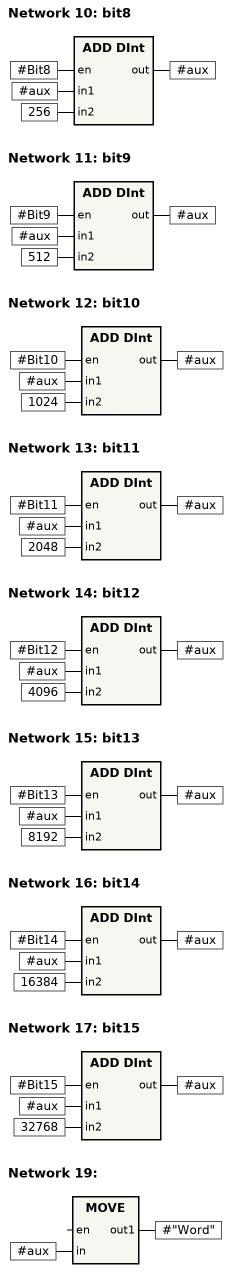
   IF #Bit8 THEN #aux := #aux + 256; END_IF;
END_REGION

REGION Network 11: bit9
   // Addiere Bit 9 zur Hilfsvariable "aux".
   // ***************************************************************************
   // Add Bit 9 to the auxiliary variable "aux".
   IF #Bit9 THEN #aux := #aux + 512; END_IF;
END_REGION

REGION Network 12: bit10
   // Addiere Bit 10 zur Hilfsvariable "aux".
   // ***************************************************************************
   // Add Bit 10 to the auxiliary variable "aux".
   IF #Bit10 THEN #aux := #aux + 1024; END_IF;
END_REGION

REGION Network 13: bit11
   // Addiere Bit 11 zur Hilfsvariable "aux".
   // ***************************************************************************
   // Add Bit 11 to the auxiliary variable "aux".
   IF #Bit11 THEN #aux := #aux + 2048; END_IF;
END_REGION

REGION Network 14: bit12
   // Addiere Bit 12 zur Hilfsvariable "aux".
   // ***************************************************************************
   // Add Bit 12 to the auxiliary variable "aux".
   IF #Bit12 THEN #aux := #aux + 4096; END_IF;
END_REGION

REGION Network 15: bit13
   // Addiere Bit 13 zur Hilfsvariable "aux".
   // ***************************************************************************
   // Add Bit 13 to the auxiliary variable "aux".
   IF #Bit13 THEN #aux := #aux + 8192; END_IF;
END_REGION

REGION Network 16: bit14
   // Addiere Bit 14 zur Hilfsvariable "aux".
   // ***************************************************************************
   // Add Bit 14 to the auxiliary variable "aux".
   IF #Bit14 THEN #aux := #aux + 16384; END_IF;
END_REGION

REGION Network 17: bit15
   // Addiere Bit 15 zur Hilfsvariable "aux".
   // ***************************************************************************
   // Add Bit 15 to the auxiliary variable "aux".
   IF #Bit15 THEN #aux := #aux + 32768; END_IF;
END_REGION

REGION Network 18: Word
   // Der Wert der Variablen "aux" wird  vom Datentyp "UInt" zum Datentyp "Word" konvertiert und der Ausgangsvariablen "Word" übergeben.
   // ***************************************************************************
   // The value of the variable "aux" will convert from type of data "UInt" to type of data "Word" and transfered to the output variable "Word".
END_REGION

REGION Network 19
   #"Word" := #aux;
END_REGION
END_FUNCTION

// folder: 60 - 69 Alarm & Satus Handling

FUNCTION "60_Alarms" : Void   // FC60, LAD
TITLE = Alarm Processing
{ S7_Optimized_Access := 'TRUE' }
AUTHOR : JRS
VERSION : 0.1
// To determine alarm conditions
   VAR_TEMP   // added for the SCL form of the ladder/FBD networks
      _w1 : Bool;
      _w2 : Bool;
   END_VAR
BEGIN

REGION Network 1: DB60 DBX0.0 = Master PLC Heart Beat Missing
   // BC_ALARM_WORD_01_BIT_0
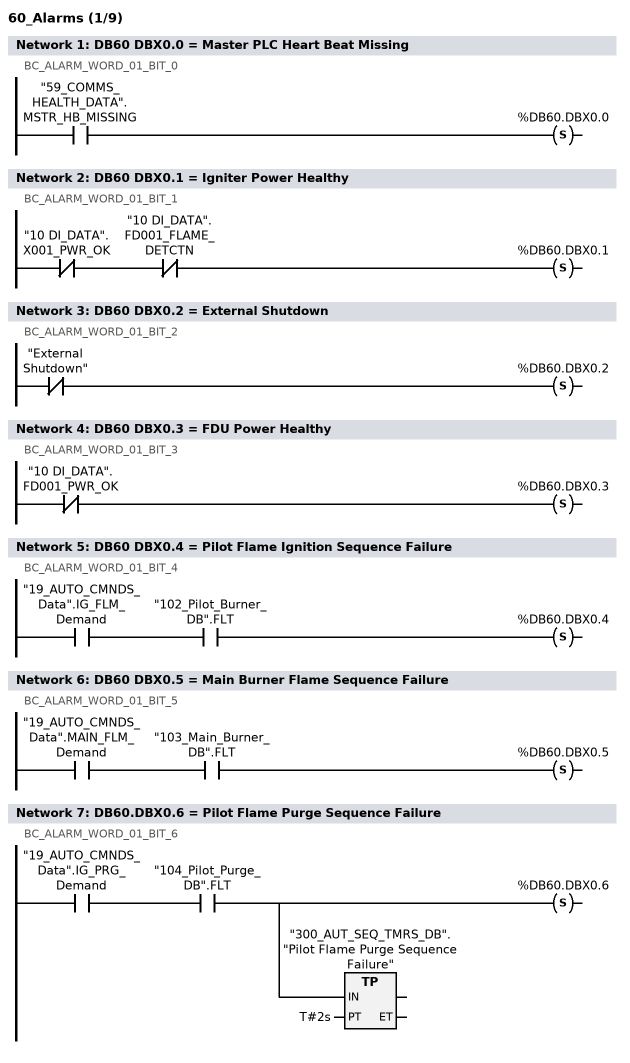
   RUNG wire#powerrail
      Contact( "59_COMMS_HEALTH_DATA".MSTR_HB_MISSING )
      S_Coil( %DB60.DBX0.0 )
   END_RUNG
   // the same network as SCL:
   IF "59_COMMS_HEALTH_DATA".MSTR_HB_MISSING THEN %DB60.DBX0.0 := TRUE; END_IF;
END_REGION

REGION Network 2: DB60 DBX0.1 = Igniter Power Healthy
   // BC_ALARM_WORD_01_BIT_1
   RUNG wire#powerrail
      I_Contact( "10 DI_DATA".X001_PWR_OK )
      I_Contact( "10 DI_DATA".FD001_FLAME_DETCTN )
      S_Coil( %DB60.DBX0.1 )
   END_RUNG
   // the same network as SCL:
   IF NOT "10 DI_DATA".X001_PWR_OK AND NOT "10 DI_DATA".FD001_FLAME_DETCTN THEN %DB60.DBX0.1 := TRUE; END_IF;
END_REGION

REGION Network 3: DB60 DBX0.2 = External Shutdown
   // BC_ALARM_WORD_01_BIT_2
   RUNG wire#powerrail
      I_Contact( "External Shutdown" )
      S_Coil( %DB60.DBX0.2 )
   END_RUNG
   // the same network as SCL:
   IF NOT "External Shutdown" THEN %DB60.DBX0.2 := TRUE; END_IF;
END_REGION

REGION Network 4: DB60 DBX0.3 = FDU Power Healthy
   // BC_ALARM_WORD_01_BIT_3
   RUNG wire#powerrail
      I_Contact( "10 DI_DATA".FD001_PWR_OK )
      S_Coil( %DB60.DBX0.3 )
   END_RUNG
   // the same network as SCL:
   IF NOT "10 DI_DATA".FD001_PWR_OK THEN %DB60.DBX0.3 := TRUE; END_IF;
END_REGION

REGION Network 5: DB60 DBX0.4 = Pilot Flame Ignition Sequence Failure
   // BC_ALARM_WORD_01_BIT_4
   RUNG wire#powerrail
      Contact( "19_AUTO_CMNDS_Data".IG_FLM_Demand )
      Contact( "102_Pilot_Burner_DB".FLT )
      S_Coil( %DB60.DBX0.4 )
   END_RUNG
   // the same network as SCL:
   IF "19_AUTO_CMNDS_Data".IG_FLM_Demand AND "102_Pilot_Burner_DB".FLT THEN %DB60.DBX0.4 := TRUE; END_IF;
END_REGION

REGION Network 6: DB60 DBX0.5 = Main Burner Flame Sequence Failure
   // BC_ALARM_WORD_01_BIT_5
   RUNG wire#powerrail
      Contact( "19_AUTO_CMNDS_Data".MAIN_FLM_Demand )
      Contact( "103_Main_Burner_DB".FLT )
      S_Coil( %DB60.DBX0.5 )
   END_RUNG
   // the same network as SCL:
   IF "19_AUTO_CMNDS_Data".MAIN_FLM_Demand AND "103_Main_Burner_DB".FLT THEN %DB60.DBX0.5 := TRUE; END_IF;
END_REGION

REGION Network 7: DB60.DBX0.6 = Pilot Flame Purge Sequence Failure
   // BC_ALARM_WORD_01_BIT_6
   #_w1 := "19_AUTO_CMNDS_Data".IG_PRG_Demand AND "104_Pilot_Purge_DB".FLT;
   IF #_w1 THEN %DB60.DBX0.6 := TRUE; END_IF;
   "300_AUT_SEQ_TMRS_DB"."Pilot Flame Purge Sequence Failure".TP(IN := #_w1, PT := T#2s);
END_REGION

REGION Network 8: DB60.DBX0.7 = FDU Healthy
   // BC_ALARM_WORD_01_BIT_7
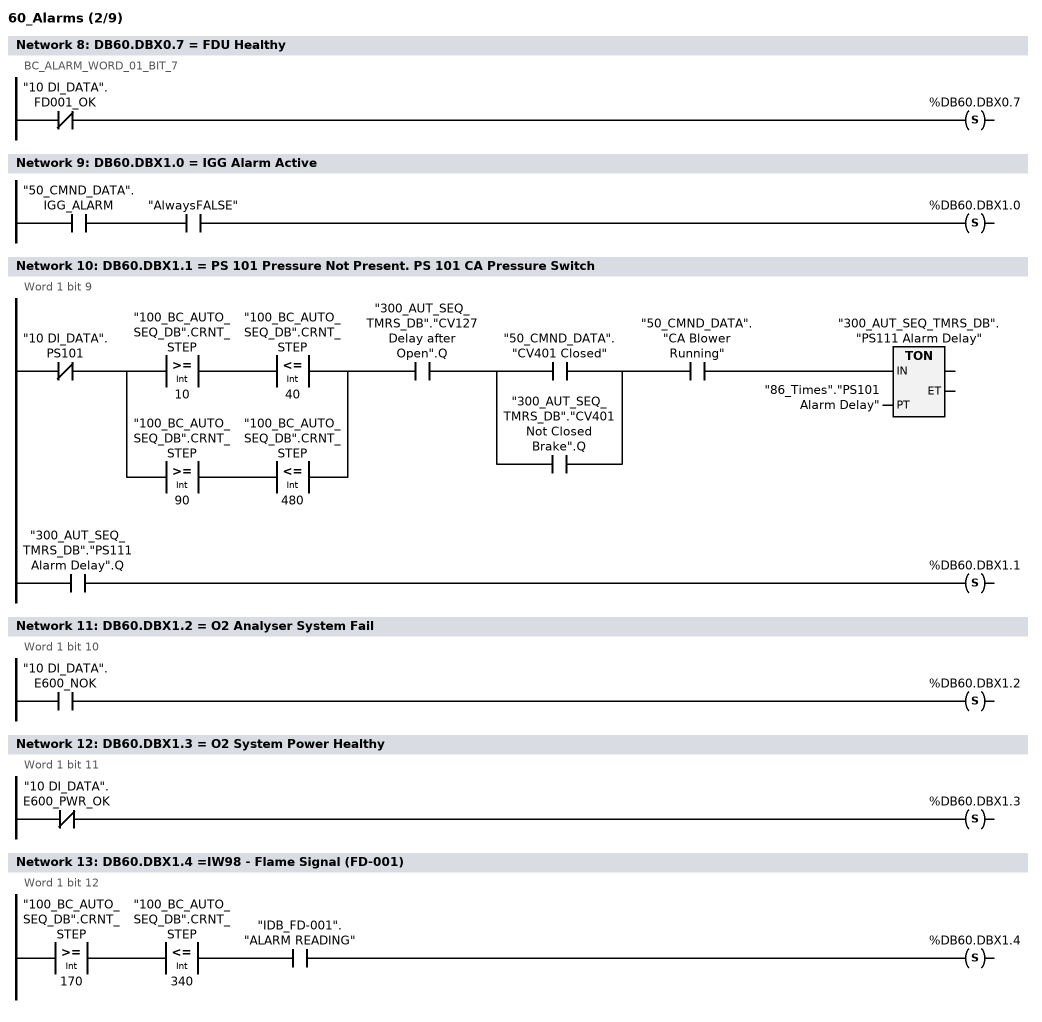
   RUNG wire#powerrail
      I_Contact( "10 DI_DATA".FD001_OK )
      S_Coil( %DB60.DBX0.7 )
   END_RUNG
   // the same network as SCL:
   IF NOT "10 DI_DATA".FD001_OK THEN %DB60.DBX0.7 := TRUE; END_IF;
END_REGION

REGION Network 9: DB60.DBX1.0 = IGG Alarm Active
   RUNG wire#powerrail
      Contact( "50_CMND_DATA".IGG_ALARM )
      Contact( "AlwaysFALSE" )
      S_Coil( %DB60.DBX1.0 )
   END_RUNG
   // the same network as SCL:
   IF "50_CMND_DATA".IGG_ALARM AND "AlwaysFALSE" THEN %DB60.DBX1.0 := TRUE; END_IF;
END_REGION

REGION Network 10: DB60.DBX1.1 = PS 101 Pressure Not Present. PS 101 CA Pressure Switch
   // Word 1 bit 9
   "300_AUT_SEQ_TMRS_DB"."PS111 Alarm Delay".TON(IN := NOT "10 DI_DATA".PS101 AND ((("100_BC_AUTO_SEQ_DB".CRNT_STEP >= 10) AND ("100_BC_AUTO_SEQ_DB".CRNT_STEP <= 40)) OR (("100_BC_AUTO_SEQ_DB".CRNT_STEP >= 90) AND ("100_BC_AUTO_SEQ_DB".CRNT_STEP <= 480))) AND "300_AUT_SEQ_TMRS_DB"."CV127 Delay after Open".Q AND ("50_CMND_DATA"."CV401 Closed" OR "300_AUT_SEQ_TMRS_DB"."CV401 Not Closed Brake".Q) AND "50_CMND_DATA"."CA Blower Running",
                           PT := "86_Times"."PS101 Alarm Delay");
   IF "300_AUT_SEQ_TMRS_DB"."PS111 Alarm Delay".Q THEN %DB60.DBX1.1 := TRUE; END_IF;
END_REGION

REGION Network 11: DB60.DBX1.2 = O2 Analyser System Fail
   // Word 1 bit 10
   RUNG wire#powerrail
      Contact( "10 DI_DATA".E600_NOK )
      S_Coil( %DB60.DBX1.2 )
   END_RUNG
   // the same network as SCL:
   IF "10 DI_DATA".E600_NOK THEN %DB60.DBX1.2 := TRUE; END_IF;
END_REGION

REGION Network 12: DB60.DBX1.3 = O2 System Power Healthy
   // Word 1 bit 11
   RUNG wire#powerrail
      I_Contact( "10 DI_DATA".E600_PWR_OK )
      S_Coil( %DB60.DBX1.3 )
   END_RUNG
   // the same network as SCL:
   IF NOT "10 DI_DATA".E600_PWR_OK THEN %DB60.DBX1.3 := TRUE; END_IF;
END_REGION

REGION Network 13: DB60.DBX1.4 =IW98 - Flame Signal (FD-001)
   // Word 1 bit 12
   RUNG wire#powerrail
      { S7_Templates := "SrcType := Int" } GE_Contact(in1 := "100_BC_AUTO_SEQ_DB".CRNT_STEP, in2 := 170)
      { S7_Templates := "SrcType := Int" } LE_Contact(in1 := "100_BC_AUTO_SEQ_DB".CRNT_STEP, in2 := 340)
      Contact( "IDB_FD-001"."ALARM READING" )
      S_Coil( %DB60.DBX1.4 )
   END_RUNG
   // the same network as SCL:
   IF ("100_BC_AUTO_SEQ_DB".CRNT_STEP >= 170) AND ("100_BC_AUTO_SEQ_DB".CRNT_STEP <= 340) AND "IDB_FD-001"."ALARM READING" THEN
       %DB60.DBX1.4 := TRUE;
   END_IF;
END_REGION

REGION Network 14: DB60.DBX1.5 =IW108 - O2 Analyser Content (E-600)
   // BC_ALARM_WORD_01 bit 13&14
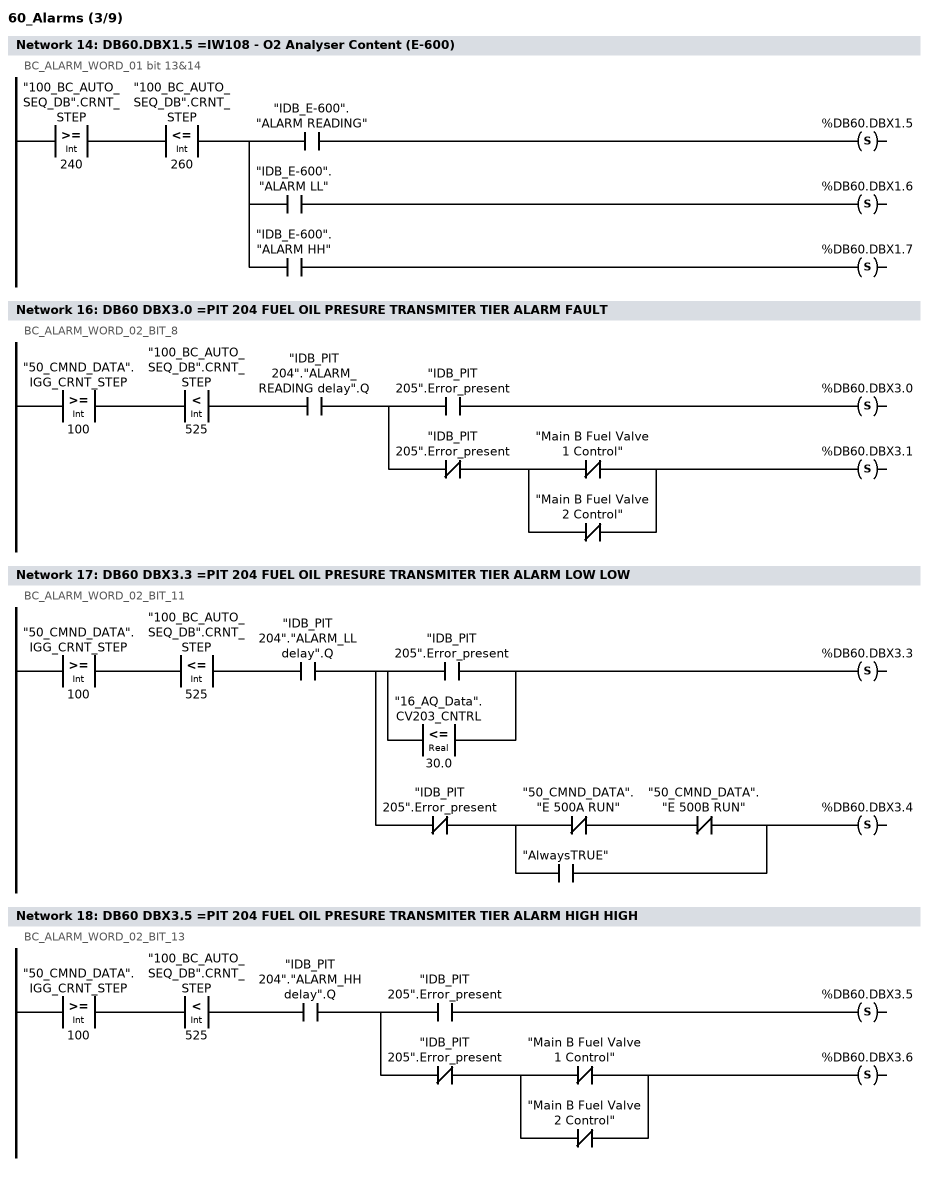
   RUNG wire#powerrail
      { S7_Templates := "SrcType := Int" } GE_Contact(in1 := "100_BC_AUTO_SEQ_DB".CRNT_STEP, in2 := 240)
      { S7_Templates := "SrcType := Int" } LE_Contact(in1 := "100_BC_AUTO_SEQ_DB".CRNT_STEP, in2 := 260)
      wire#w1
      Contact( "IDB_E-600"."ALARM READING" )
      S_Coil( %DB60.DBX1.5 )
   END_RUNG
   RUNG wire#w1
      Contact( "IDB_E-600"."ALARM LL" )
      S_Coil( %DB60.DBX1.6 )
   END_RUNG
   RUNG wire#w1
      Contact( "IDB_E-600"."ALARM HH" )
      S_Coil( %DB60.DBX1.7 )
   END_RUNG
   // the same network as SCL:
   #_w1 := ("100_BC_AUTO_SEQ_DB".CRNT_STEP >= 240) AND ("100_BC_AUTO_SEQ_DB".CRNT_STEP <= 260);
   IF #_w1 AND "IDB_E-600"."ALARM READING" THEN %DB60.DBX1.5 := TRUE; END_IF;
   IF #_w1 AND "IDB_E-600"."ALARM LL" THEN %DB60.DBX1.6 := TRUE; END_IF;
   IF #_w1 AND "IDB_E-600"."ALARM HH" THEN %DB60.DBX1.7 := TRUE; END_IF;
END_REGION

REGION Network 16: DB60 DBX3.0 =PIT 204 FUEL OIL PRESURE TRANSMITER TIER ALARM FAULT
   // BC_ALARM_WORD_02_BIT_8
   RUNG wire#powerrail
      { S7_Templates := "SrcType := Int" } GE_Contact(in1 := "50_CMND_DATA".IGG_CRNT_STEP, in2 := 100)
      { S7_Templates := "SrcType := Int" } LT_Contact(in1 := "100_BC_AUTO_SEQ_DB".CRNT_STEP, in2 := 525)
      Contact( "IDB_PIT 204"."ALARM_READING delay".Q )
      wire#w1
      Contact( "IDB_PIT 205".Error_present )
      S_Coil( %DB60.DBX3.0 )
   END_RUNG
   RUNG wire#w1
      I_Contact( "IDB_PIT 205".Error_present )
      wire#w2
      I_Contact( "Main B Fuel Valve 1 Control" )
      wire#w3
      S_Coil( %DB60.DBX3.1 )
   END_RUNG
   RUNG wire#w2
      I_Contact( "Main B Fuel Valve 2 Control" )
   END_RUNG wire#w3
   // the same network as SCL:
   #_w1 := ("50_CMND_DATA".IGG_CRNT_STEP >= 100) AND ("100_BC_AUTO_SEQ_DB".CRNT_STEP < 525) AND "IDB_PIT 204"."ALARM_READING delay".Q;
   IF #_w1 AND "IDB_PIT 205".Error_present THEN %DB60.DBX3.0 := TRUE; END_IF;
   IF #_w1 AND NOT "IDB_PIT 205".Error_present AND (NOT "Main B Fuel Valve 1 Control" OR NOT "Main B Fuel Valve 2 Control") THEN
       %DB60.DBX3.1 := TRUE;
   END_IF;
END_REGION

REGION Network 17: DB60 DBX3.3 =PIT 204 FUEL OIL PRESURE TRANSMITER TIER ALARM LOW LOW
   // BC_ALARM_WORD_02_BIT_11
   RUNG wire#powerrail
      { S7_Templates := "SrcType := Int" } GE_Contact(in1 := "50_CMND_DATA".IGG_CRNT_STEP, in2 := 100)
      { S7_Templates := "SrcType := Int" } LE_Contact(in1 := "100_BC_AUTO_SEQ_DB".CRNT_STEP, in2 := 525)
      Contact( "IDB_PIT 204"."ALARM_LL delay".Q )
      wire#w1
      Contact( "IDB_PIT 205".Error_present )
      wire#w2
      S_Coil( %DB60.DBX3.3 )
   END_RUNG
   RUNG wire#w1
      { S7_Templates := "SrcType := Real" } LE_Contact(in1 := "16_AQ_Data".CV203_CNTRL, in2 := 30.0)
   END_RUNG wire#w2
   RUNG wire#w1
      I_Contact( "IDB_PIT 205".Error_present )
      wire#w3
      I_Contact( "50_CMND_DATA"."E 500A RUN" )
      I_Contact( "50_CMND_DATA"."E 500B RUN" )
      wire#w4
      S_Coil( %DB60.DBX3.4 )
   END_RUNG
   RUNG wire#w3
      Contact( "AlwaysTRUE" )
   END_RUNG wire#w4
   // the same network as SCL:
   #_w1 := ("50_CMND_DATA".IGG_CRNT_STEP >= 100) AND ("100_BC_AUTO_SEQ_DB".CRNT_STEP <= 525) AND "IDB_PIT 204"."ALARM_LL delay".Q;
   IF #_w1 AND ("IDB_PIT 205".Error_present OR ("16_AQ_Data".CV203_CNTRL <= 30.0)) THEN
       %DB60.DBX3.3 := TRUE;
   END_IF;
   IF #_w1 AND NOT "IDB_PIT 205".Error_present AND ((NOT "50_CMND_DATA"."E 500A RUN" AND NOT "50_CMND_DATA"."E 500B RUN") OR "AlwaysTRUE") THEN
       %DB60.DBX3.4 := TRUE;
   END_IF;
END_REGION

REGION Network 18: DB60 DBX3.5 =PIT 204 FUEL OIL PRESURE TRANSMITER TIER ALARM HIGH HIGH
   // BC_ALARM_WORD_02_BIT_13
   RUNG wire#powerrail
      { S7_Templates := "SrcType := Int" } GE_Contact(in1 := "50_CMND_DATA".IGG_CRNT_STEP, in2 := 100)
      { S7_Templates := "SrcType := Int" } LT_Contact(in1 := "100_BC_AUTO_SEQ_DB".CRNT_STEP, in2 := 525)
      Contact( "IDB_PIT 204"."ALARM_HH delay".Q )
      wire#w1
      Contact( "IDB_PIT 205".Error_present )
      S_Coil( %DB60.DBX3.5 )
   END_RUNG
   RUNG wire#w1
      I_Contact( "IDB_PIT 205".Error_present )
      wire#w2
      I_Contact( "Main B Fuel Valve 1 Control" )
      wire#w3
      S_Coil( %DB60.DBX3.6 )
   END_RUNG
   RUNG wire#w2
      I_Contact( "Main B Fuel Valve 2 Control" )
   END_RUNG wire#w3
   // the same network as SCL:
   #_w1 := ("50_CMND_DATA".IGG_CRNT_STEP >= 100) AND ("100_BC_AUTO_SEQ_DB".CRNT_STEP < 525) AND "IDB_PIT 204"."ALARM_HH delay".Q;
   IF #_w1 AND "IDB_PIT 205".Error_present THEN %DB60.DBX3.5 := TRUE; END_IF;
   IF #_w1 AND NOT "IDB_PIT 205".Error_present AND (NOT "Main B Fuel Valve 1 Control" OR NOT "Main B Fuel Valve 2 Control") THEN
       %DB60.DBX3.6 := TRUE;
   END_IF;
END_REGION

REGION Network 19: DB60 DBX4.0 =FS 123 PILOT BURNER AIR FLOW SWITCH
   // BC_ALARM_WORD_03_BIT_0
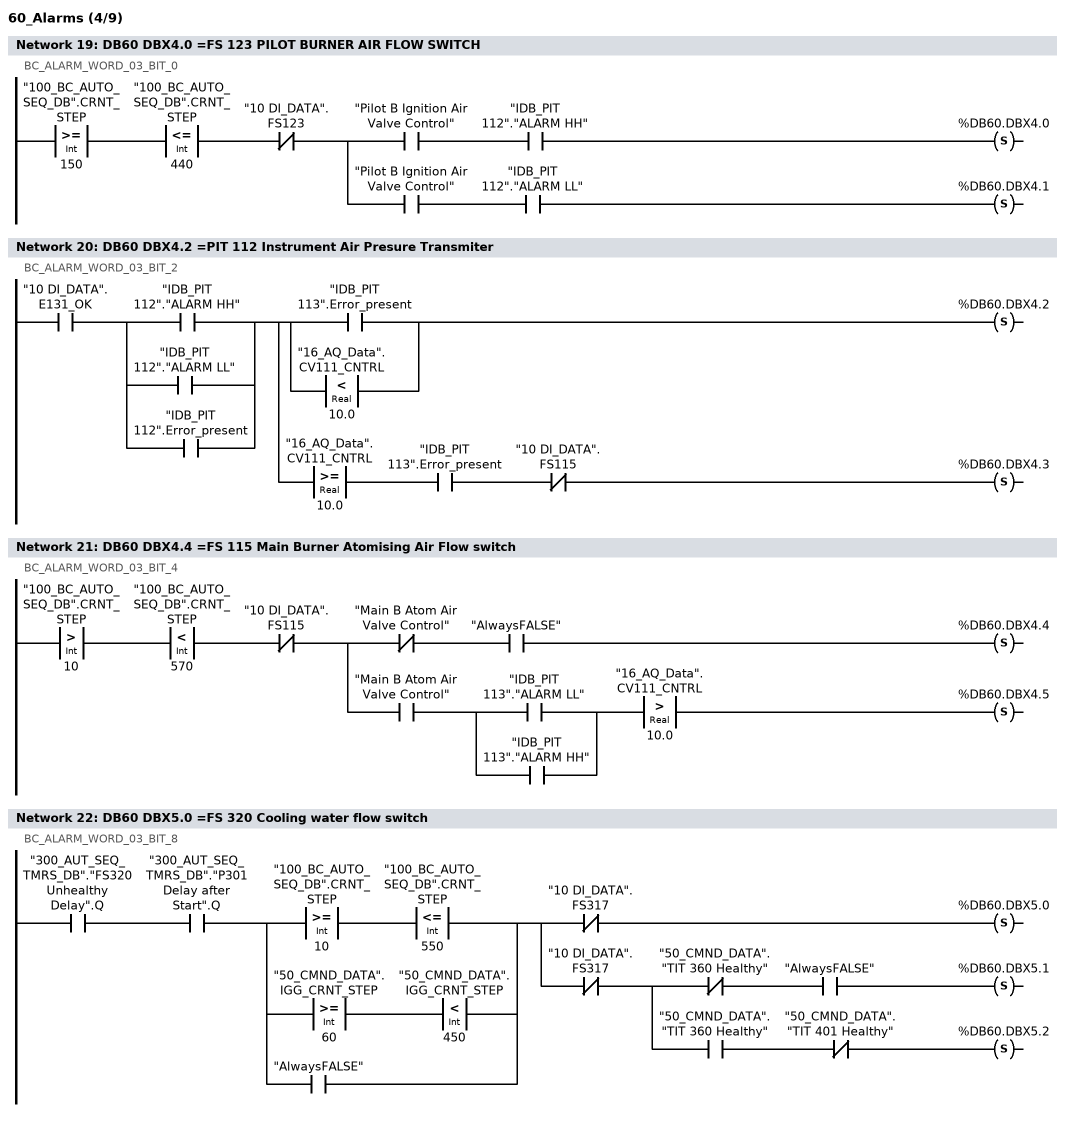
   RUNG wire#powerrail
      { S7_Templates := "SrcType := Int" } GE_Contact(in1 := "100_BC_AUTO_SEQ_DB".CRNT_STEP, in2 := 150)
      { S7_Templates := "SrcType := Int" } LE_Contact(in1 := "100_BC_AUTO_SEQ_DB".CRNT_STEP, in2 := 440)
      I_Contact( "10 DI_DATA".FS123 )
      wire#w1
      Contact( "Pilot B Ignition Air Valve Control" )
      Contact( "IDB_PIT 112"."ALARM HH" )
      S_Coil( %DB60.DBX4.0 )
   END_RUNG
   RUNG wire#w1
      Contact( "Pilot B Ignition Air Valve Control" )
      Contact( "IDB_PIT 112"."ALARM LL" )
      S_Coil( %DB60.DBX4.1 )
   END_RUNG
   // the same network as SCL:
   #_w1 := ("100_BC_AUTO_SEQ_DB".CRNT_STEP >= 150) AND ("100_BC_AUTO_SEQ_DB".CRNT_STEP <= 440) AND NOT "10 DI_DATA".FS123;
   IF #_w1 AND "Pilot B Ignition Air Valve Control" AND "IDB_PIT 112"."ALARM HH" THEN
       %DB60.DBX4.0 := TRUE;
   END_IF;
   IF #_w1 AND "Pilot B Ignition Air Valve Control" AND "IDB_PIT 112"."ALARM LL" THEN
       %DB60.DBX4.1 := TRUE;
   END_IF;
END_REGION

REGION Network 20: DB60 DBX4.2 =PIT 112 Instrument Air Presure Transmiter
   // BC_ALARM_WORD_03_BIT_2
   RUNG wire#powerrail
      Contact( "10 DI_DATA".E131_OK )
      wire#w1
      Contact( "IDB_PIT 112"."ALARM HH" )
      wire#w2
      Contact( "IDB_PIT 113".Error_present )
      wire#w3
      S_Coil( %DB60.DBX4.2 )
   END_RUNG
   RUNG wire#w1
      Contact( "IDB_PIT 112"."ALARM LL" )
   END_RUNG wire#w2
   RUNG wire#w1
      Contact( "IDB_PIT 112".Error_present )
   END_RUNG wire#w2
   RUNG wire#w2
      { S7_Templates := "SrcType := Real" } LT_Contact(in1 := "16_AQ_Data".CV111_CNTRL, in2 := 10.0)
   END_RUNG wire#w3
   RUNG wire#w2
      { S7_Templates := "SrcType := Real" } GE_Contact(in1 := "16_AQ_Data".CV111_CNTRL, in2 := 10.0)
      Contact( "IDB_PIT 113".Error_present )
      I_Contact( "10 DI_DATA".FS115 )
      S_Coil( %DB60.DBX4.3 )
   END_RUNG
   // the same network as SCL:
   #_w1 := "10 DI_DATA".E131_OK AND ("IDB_PIT 112"."ALARM HH" OR "IDB_PIT 112"."ALARM LL" OR "IDB_PIT 112".Error_present);
   IF #_w1 AND ("IDB_PIT 113".Error_present OR ("16_AQ_Data".CV111_CNTRL < 10.0)) THEN
       %DB60.DBX4.2 := TRUE;
   END_IF;
   IF #_w1 AND ("16_AQ_Data".CV111_CNTRL >= 10.0) AND "IDB_PIT 113".Error_present AND NOT "10 DI_DATA".FS115 THEN
       %DB60.DBX4.3 := TRUE;
   END_IF;
END_REGION

REGION Network 21: DB60 DBX4.4 =FS 115 Main Burner Atomising Air Flow switch
   // BC_ALARM_WORD_03_BIT_4
   RUNG wire#powerrail
      { S7_Templates := "SrcType := Int" } GT_Contact(in1 := "100_BC_AUTO_SEQ_DB".CRNT_STEP, in2 := 10)
      { S7_Templates := "SrcType := Int" } LT_Contact(in1 := "100_BC_AUTO_SEQ_DB".CRNT_STEP, in2 := 570)
      I_Contact( "10 DI_DATA".FS115 )
      wire#w1
      I_Contact( "Main B Atom Air Valve Control" )
      Contact( "AlwaysFALSE" )
      S_Coil( %DB60.DBX4.4 )
   END_RUNG
   RUNG wire#w1
      Contact( "Main B Atom Air Valve Control" )
      wire#w2
      Contact( "IDB_PIT 113"."ALARM LL" )
      wire#w3
      { S7_Templates := "SrcType := Real" } GT_Contact(in1 := "16_AQ_Data".CV111_CNTRL, in2 := 10.0)
      S_Coil( %DB60.DBX4.5 )
   END_RUNG
   RUNG wire#w2
      Contact( "IDB_PIT 113"."ALARM HH" )
   END_RUNG wire#w3
   // the same network as SCL:
   #_w1 := ("100_BC_AUTO_SEQ_DB".CRNT_STEP > 10) AND ("100_BC_AUTO_SEQ_DB".CRNT_STEP < 570) AND NOT "10 DI_DATA".FS115;
   IF #_w1 AND NOT "Main B Atom Air Valve Control" AND "AlwaysFALSE" THEN %DB60.DBX4.4 := TRUE; END_IF;
   IF #_w1 AND "Main B Atom Air Valve Control" AND ("IDB_PIT 113"."ALARM LL" OR "IDB_PIT 113"."ALARM HH") AND ("16_AQ_Data".CV111_CNTRL > 10.0) THEN
       %DB60.DBX4.5 := TRUE;
   END_IF;
END_REGION

REGION Network 22: DB60 DBX5.0 =FS 320 Cooling water flow switch
   // BC_ALARM_WORD_03_BIT_8
   RUNG wire#powerrail
      Contact( "300_AUT_SEQ_TMRS_DB"."FS320 Unhealthy Delay".Q )
      Contact( "300_AUT_SEQ_TMRS_DB"."P301 Delay after Start".Q )
      wire#w1
      { S7_Templates := "SrcType := Int" } GE_Contact(in1 := "100_BC_AUTO_SEQ_DB".CRNT_STEP, in2 := 10)
      { S7_Templates := "SrcType := Int" } LE_Contact(in1 := "100_BC_AUTO_SEQ_DB".CRNT_STEP, in2 := 550)
      wire#w2
      I_Contact( "10 DI_DATA".FS317 )
      S_Coil( %DB60.DBX5.0 )
   END_RUNG
   RUNG wire#w1
      { S7_Templates := "SrcType := Int" } GE_Contact(in1 := "50_CMND_DATA".IGG_CRNT_STEP, in2 := 60)
      { S7_Templates := "SrcType := Int" } LT_Contact(in1 := "50_CMND_DATA".IGG_CRNT_STEP, in2 := 450)
   END_RUNG wire#w2
   RUNG wire#w1
      Contact( "AlwaysFALSE" )
   END_RUNG wire#w2
   RUNG wire#w2
      I_Contact( "10 DI_DATA".FS317 )
      wire#w3
      I_Contact( "50_CMND_DATA"."TIT 360 Healthy" )
      Contact( "AlwaysFALSE" )
      S_Coil( %DB60.DBX5.1 )
   END_RUNG
   RUNG wire#w3
      Contact( "50_CMND_DATA"."TIT 360 Healthy" )
      I_Contact( "50_CMND_DATA"."TIT 401 Healthy" )
      S_Coil( %DB60.DBX5.2 )
   END_RUNG
   // the same network as SCL:
   #_w1 := "300_AUT_SEQ_TMRS_DB"."FS320 Unhealthy Delay".Q AND "300_AUT_SEQ_TMRS_DB"."P301 Delay after Start".Q AND ((("100_BC_AUTO_SEQ_DB".CRNT_STEP >= 10) AND ("100_BC_AUTO_SEQ_DB".CRNT_STEP <= 550)) OR (("50_CMND_DATA".IGG_CRNT_STEP >= 60) AND ("50_CMND_DATA".IGG_CRNT_STEP < 450)) OR "AlwaysFALSE");
   IF #_w1 AND NOT "10 DI_DATA".FS317 THEN %DB60.DBX5.0 := TRUE; END_IF;
   #_w2 := #_w1 AND NOT "10 DI_DATA".FS317;
   IF #_w2 AND NOT "50_CMND_DATA"."TIT 360 Healthy" AND "AlwaysFALSE" THEN %DB60.DBX5.1 := TRUE; END_IF;
   IF #_w2 AND "50_CMND_DATA"."TIT 360 Healthy" AND NOT "50_CMND_DATA"."TIT 401 Healthy" THEN
       %DB60.DBX5.2 := TRUE;
   END_IF;
END_REGION

REGION Network 23: DB60 DBX5.3 =FS 317 Jacket Cooling Water Flow Switch
   // BC_ALARM_WORD_03_BIT_11
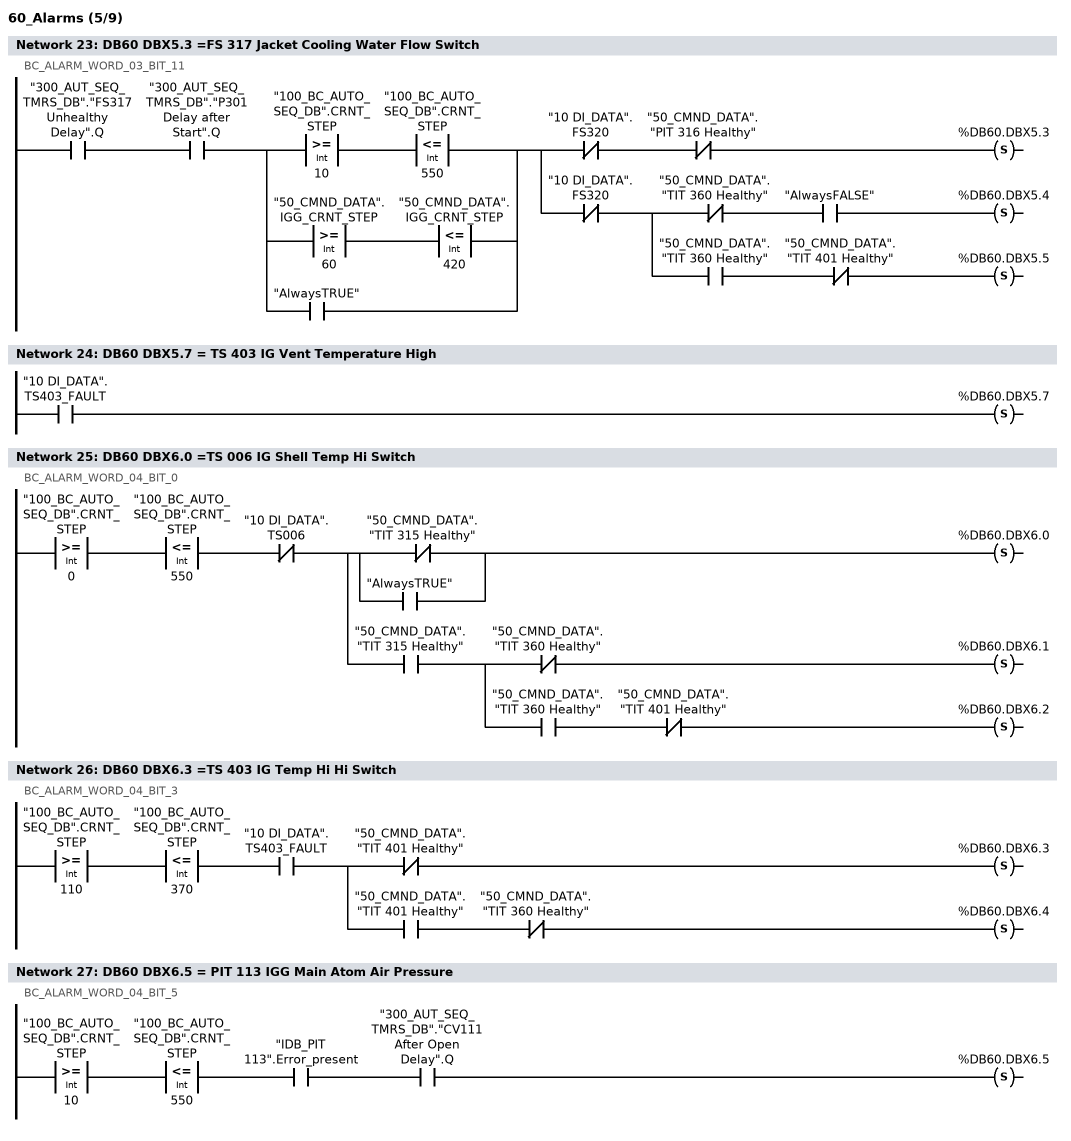
   RUNG wire#powerrail
      Contact( "300_AUT_SEQ_TMRS_DB"."FS317 Unhealthy Delay".Q )
      Contact( "300_AUT_SEQ_TMRS_DB"."P301 Delay after Start".Q )
      wire#w1
      { S7_Templates := "SrcType := Int" } GE_Contact(in1 := "100_BC_AUTO_SEQ_DB".CRNT_STEP, in2 := 10)
      { S7_Templates := "SrcType := Int" } LE_Contact(in1 := "100_BC_AUTO_SEQ_DB".CRNT_STEP, in2 := 550)
      wire#w2
      I_Contact( "10 DI_DATA".FS320 )
      I_Contact( "50_CMND_DATA"."PIT 316 Healthy" )
      S_Coil( %DB60.DBX5.3 )
   END_RUNG
   RUNG wire#w1
      { S7_Templates := "SrcType := Int" } GE_Contact(in1 := "50_CMND_DATA".IGG_CRNT_STEP, in2 := 60)
      { S7_Templates := "SrcType := Int" } LE_Contact(in1 := "50_CMND_DATA".IGG_CRNT_STEP, in2 := 420)
   END_RUNG wire#w2
   RUNG wire#w1
      Contact( "AlwaysTRUE" )
   END_RUNG wire#w2
   RUNG wire#w2
      I_Contact( "10 DI_DATA".FS320 )
      wire#w3
      I_Contact( "50_CMND_DATA"."TIT 360 Healthy" )
      Contact( "AlwaysFALSE" )
      S_Coil( %DB60.DBX5.4 )
   END_RUNG
   RUNG wire#w3
      Contact( "50_CMND_DATA"."TIT 360 Healthy" )
      I_Contact( "50_CMND_DATA"."TIT 401 Healthy" )
      S_Coil( %DB60.DBX5.5 )
   END_RUNG
   // the same network as SCL:
   #_w1 := "300_AUT_SEQ_TMRS_DB"."FS317 Unhealthy Delay".Q AND "300_AUT_SEQ_TMRS_DB"."P301 Delay after Start".Q AND ((("100_BC_AUTO_SEQ_DB".CRNT_STEP >= 10) AND ("100_BC_AUTO_SEQ_DB".CRNT_STEP <= 550)) OR (("50_CMND_DATA".IGG_CRNT_STEP >= 60) AND ("50_CMND_DATA".IGG_CRNT_STEP <= 420)) OR "AlwaysTRUE");
   IF #_w1 AND NOT "10 DI_DATA".FS320 AND NOT "50_CMND_DATA"."PIT 316 Healthy" THEN
       %DB60.DBX5.3 := TRUE;
   END_IF;
   #_w2 := #_w1 AND NOT "10 DI_DATA".FS320;
   IF #_w2 AND NOT "50_CMND_DATA"."TIT 360 Healthy" AND "AlwaysFALSE" THEN %DB60.DBX5.4 := TRUE; END_IF;
   IF #_w2 AND "50_CMND_DATA"."TIT 360 Healthy" AND NOT "50_CMND_DATA"."TIT 401 Healthy" THEN
       %DB60.DBX5.5 := TRUE;
   END_IF;
END_REGION

REGION Network 24: DB60 DBX5.7 = TS 403 IG Vent Temperature High
   RUNG wire#powerrail
      Contact( "10 DI_DATA".TS403_FAULT )
      S_Coil( %DB60.DBX5.7 )
   END_RUNG
   // the same network as SCL:
   IF "10 DI_DATA".TS403_FAULT THEN %DB60.DBX5.7 := TRUE; END_IF;
END_REGION

REGION Network 25: DB60 DBX6.0 =TS 006 IG Shell Temp Hi Switch
   // BC_ALARM_WORD_04_BIT_0
   RUNG wire#powerrail
      { S7_Templates := "SrcType := Int" } GE_Contact(in1 := "100_BC_AUTO_SEQ_DB".CRNT_STEP, in2 := 0)
      { S7_Templates := "SrcType := Int" } LE_Contact(in1 := "100_BC_AUTO_SEQ_DB".CRNT_STEP, in2 := 550)
      I_Contact( "10 DI_DATA".TS006 )
      wire#w1
      I_Contact( "50_CMND_DATA"."TIT 315 Healthy" )
      wire#w2
      S_Coil( %DB60.DBX6.0 )
   END_RUNG
   RUNG wire#w1
      Contact( "AlwaysTRUE" )
   END_RUNG wire#w2
   RUNG wire#w1
      Contact( "50_CMND_DATA"."TIT 315 Healthy" )
      wire#w3
      I_Contact( "50_CMND_DATA"."TIT 360 Healthy" )
      S_Coil( %DB60.DBX6.1 )
   END_RUNG
   RUNG wire#w3
      Contact( "50_CMND_DATA"."TIT 360 Healthy" )
      I_Contact( "50_CMND_DATA"."TIT 401 Healthy" )
      S_Coil( %DB60.DBX6.2 )
   END_RUNG
   // the same network as SCL:
   #_w1 := ("100_BC_AUTO_SEQ_DB".CRNT_STEP >= 0) AND ("100_BC_AUTO_SEQ_DB".CRNT_STEP <= 550) AND NOT "10 DI_DATA".TS006;
   IF #_w1 AND (NOT "50_CMND_DATA"."TIT 315 Healthy" OR "AlwaysTRUE") THEN %DB60.DBX6.0 := TRUE; END_IF;
   #_w2 := #_w1 AND "50_CMND_DATA"."TIT 315 Healthy";
   IF #_w2 AND NOT "50_CMND_DATA"."TIT 360 Healthy" THEN %DB60.DBX6.1 := TRUE; END_IF;
   IF #_w2 AND "50_CMND_DATA"."TIT 360 Healthy" AND NOT "50_CMND_DATA"."TIT 401 Healthy" THEN
       %DB60.DBX6.2 := TRUE;
   END_IF;
END_REGION

REGION Network 26: DB60 DBX6.3 =TS 403 IG Temp Hi Hi Switch
   // BC_ALARM_WORD_04_BIT_3
   RUNG wire#powerrail
      { S7_Templates := "SrcType := Int" } GE_Contact(in1 := "100_BC_AUTO_SEQ_DB".CRNT_STEP, in2 := 110)
      { S7_Templates := "SrcType := Int" } LE_Contact(in1 := "100_BC_AUTO_SEQ_DB".CRNT_STEP, in2 := 370)
      Contact( "10 DI_DATA".TS403_FAULT )
      wire#w1
      I_Contact( "50_CMND_DATA"."TIT 401 Healthy" )
      S_Coil( %DB60.DBX6.3 )
   END_RUNG
   RUNG wire#w1
      Contact( "50_CMND_DATA"."TIT 401 Healthy" )
      I_Contact( "50_CMND_DATA"."TIT 360 Healthy" )
      S_Coil( %DB60.DBX6.4 )
   END_RUNG
   // the same network as SCL:
   #_w1 := ("100_BC_AUTO_SEQ_DB".CRNT_STEP >= 110) AND ("100_BC_AUTO_SEQ_DB".CRNT_STEP <= 370) AND "10 DI_DATA".TS403_FAULT;
   IF #_w1 AND NOT "50_CMND_DATA"."TIT 401 Healthy" THEN %DB60.DBX6.3 := TRUE; END_IF;
   IF #_w1 AND "50_CMND_DATA"."TIT 401 Healthy" AND NOT "50_CMND_DATA"."TIT 360 Healthy" THEN
       %DB60.DBX6.4 := TRUE;
   END_IF;
END_REGION

REGION Network 27: DB60 DBX6.5 = PIT 113 IGG Main Atom Air Pressure
   // BC_ALARM_WORD_04_BIT_5
   RUNG wire#powerrail
      { S7_Templates := "SrcType := Int" } GE_Contact(in1 := "100_BC_AUTO_SEQ_DB".CRNT_STEP, in2 := 10)
      { S7_Templates := "SrcType := Int" } LE_Contact(in1 := "100_BC_AUTO_SEQ_DB".CRNT_STEP, in2 := 550)
      Contact( "IDB_PIT 113".Error_present )
      Contact( "300_AUT_SEQ_TMRS_DB"."CV111 After Open Delay".Q )
      S_Coil( %DB60.DBX6.5 )
   END_RUNG
   // the same network as SCL:
   IF ("100_BC_AUTO_SEQ_DB".CRNT_STEP >= 10) AND ("100_BC_AUTO_SEQ_DB".CRNT_STEP <= 550) AND "IDB_PIT 113".Error_present AND "300_AUT_SEQ_TMRS_DB"."CV111 After Open Delay".Q THEN
       %DB60.DBX6.5 := TRUE;
   END_IF;
END_REGION

REGION Network 28: DB60 DBX6.6 = PIT 205 IGG Main Fuel Pressure
   // BC_ALARM_WORD_04_BIT_6
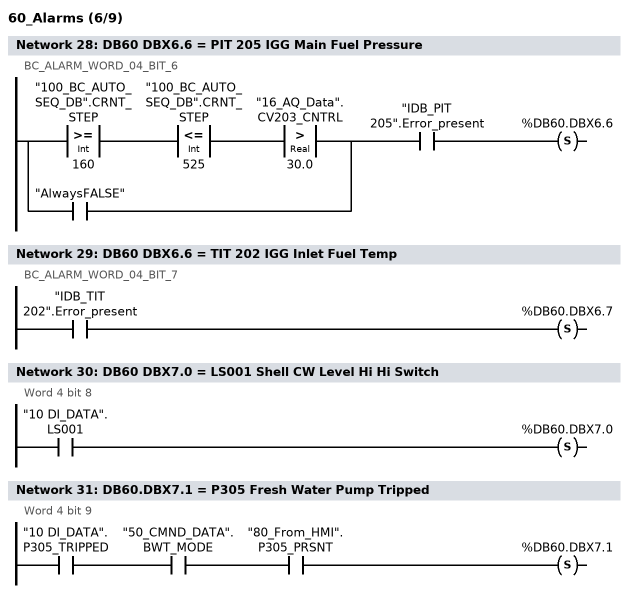
   RUNG wire#powerrail
      { S7_Templates := "SrcType := Int" } GE_Contact(in1 := "100_BC_AUTO_SEQ_DB".CRNT_STEP, in2 := 160)
      { S7_Templates := "SrcType := Int" } LE_Contact(in1 := "100_BC_AUTO_SEQ_DB".CRNT_STEP, in2 := 525)
      { S7_Templates := "SrcType := Real" } GT_Contact(in1 := "16_AQ_Data".CV203_CNTRL, in2 := 30.0)
      wire#w1
      Contact( "IDB_PIT 205".Error_present )
      S_Coil( %DB60.DBX6.6 )
   END_RUNG
   RUNG wire#powerrail
      Contact( "AlwaysFALSE" )
   END_RUNG wire#w1
   // the same network as SCL:
   IF ((("100_BC_AUTO_SEQ_DB".CRNT_STEP >= 160) AND ("100_BC_AUTO_SEQ_DB".CRNT_STEP <= 525) AND ("16_AQ_Data".CV203_CNTRL > 30.0)) OR "AlwaysFALSE") AND "IDB_PIT 205".Error_present THEN
       %DB60.DBX6.6 := TRUE;
   END_IF;
END_REGION

REGION Network 29: DB60 DBX6.6 = TIT 202 IGG Inlet Fuel Temp
   // BC_ALARM_WORD_04_BIT_7
   RUNG wire#powerrail
      Contact( "IDB_TIT 202".Error_present )
      S_Coil( %DB60.DBX6.7 )
   END_RUNG
   // the same network as SCL:
   IF "IDB_TIT 202".Error_present THEN %DB60.DBX6.7 := TRUE; END_IF;
END_REGION

REGION Network 30: DB60 DBX7.0 = LS001 Shell CW Level Hi Hi Switch
   // Word 4 bit 8
   RUNG wire#powerrail
      Contact( "10 DI_DATA".LS001 )
      S_Coil( %DB60.DBX7.0 )
   END_RUNG
   // the same network as SCL:
   IF "10 DI_DATA".LS001 THEN %DB60.DBX7.0 := TRUE; END_IF;
END_REGION

REGION Network 31: DB60.DBX7.1 = P305 Fresh Water Pump Tripped
   // Word 4 bit 9
   RUNG wire#powerrail
      Contact( "10 DI_DATA".P305_TRIPPED )
      Contact( "50_CMND_DATA".BWT_MODE )
      Contact( "80_From_HMI".P305_PRSNT )
      S_Coil( %DB60.DBX7.1 )
   END_RUNG
   // the same network as SCL:
   IF "10 DI_DATA".P305_TRIPPED AND "50_CMND_DATA".BWT_MODE AND "80_From_HMI".P305_PRSNT THEN
       %DB60.DBX7.1 := TRUE;
   END_IF;
END_REGION

REGION Network 33: Alarm reset
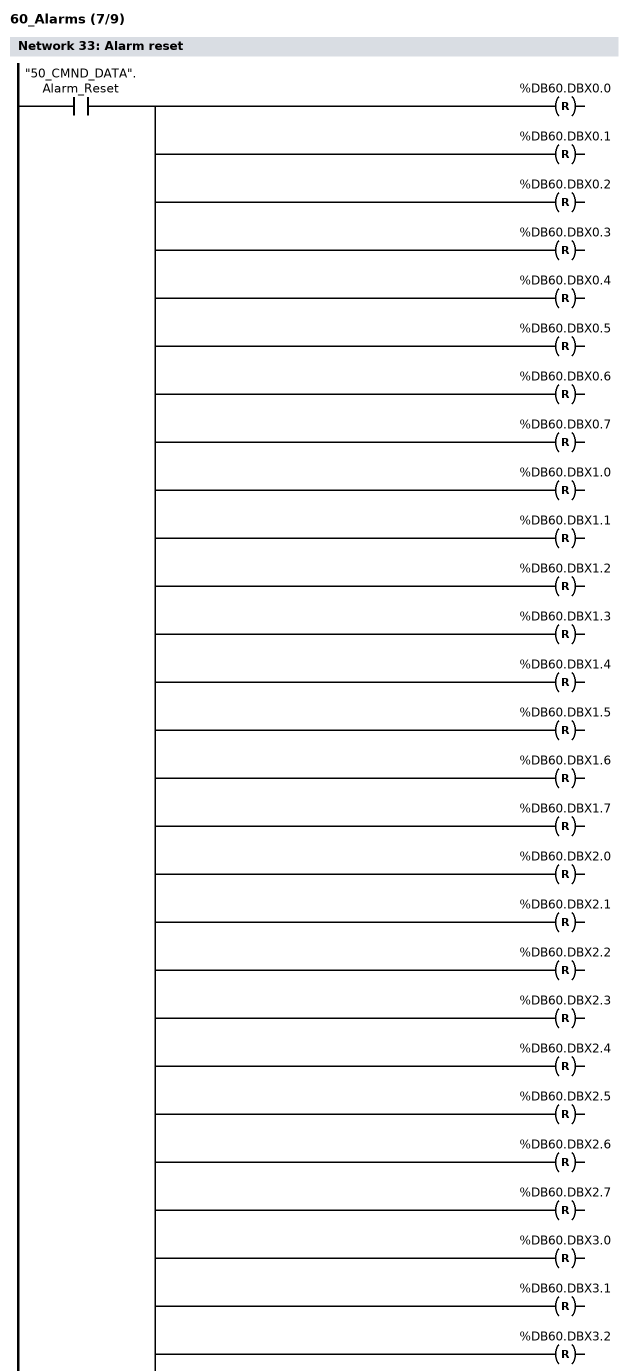
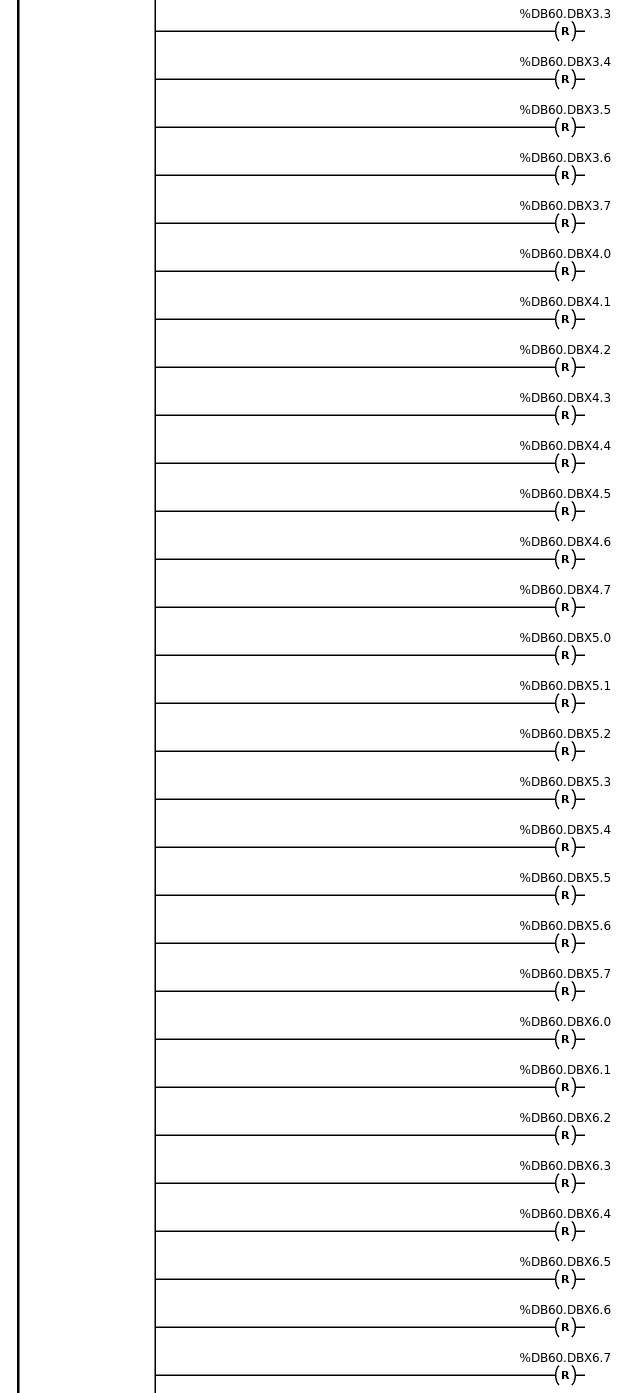
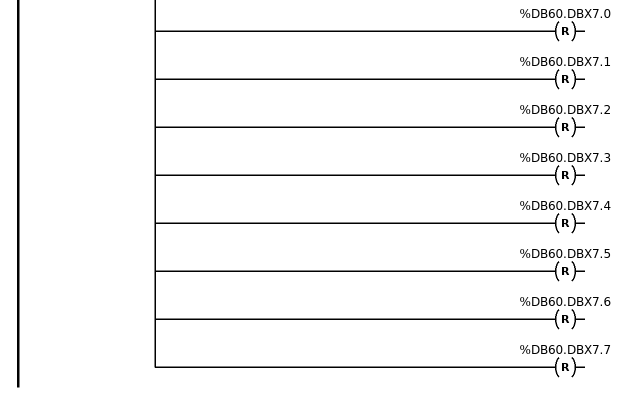
   RUNG wire#powerrail
      Contact( "50_CMND_DATA".Alarm_Reset )
      wire#w1
      R_Coil( %DB60.DBX0.0 )
   END_RUNG
   RUNG wire#w1
      R_Coil( %DB60.DBX0.1 )
   END_RUNG
   RUNG wire#w1
      R_Coil( %DB60.DBX0.2 )
   END_RUNG
   RUNG wire#w1
      R_Coil( %DB60.DBX0.3 )
   END_RUNG
   RUNG wire#w1
      R_Coil( %DB60.DBX0.4 )
   END_RUNG
   RUNG wire#w1
      R_Coil( %DB60.DBX0.5 )
   END_RUNG
   RUNG wire#w1
      R_Coil( %DB60.DBX0.6 )
   END_RUNG
   RUNG wire#w1
      R_Coil( %DB60.DBX0.7 )
   END_RUNG
   RUNG wire#w1
      R_Coil( %DB60.DBX1.0 )
   END_RUNG
   RUNG wire#w1
      R_Coil( %DB60.DBX1.1 )
   END_RUNG
   RUNG wire#w1
      R_Coil( %DB60.DBX1.2 )
   END_RUNG
   RUNG wire#w1
      R_Coil( %DB60.DBX1.3 )
   END_RUNG
   RUNG wire#w1
      R_Coil( %DB60.DBX1.4 )
   END_RUNG
   RUNG wire#w1
      R_Coil( %DB60.DBX1.5 )
   END_RUNG
   RUNG wire#w1
      R_Coil( %DB60.DBX1.6 )
   END_RUNG
   RUNG wire#w1
      R_Coil( %DB60.DBX1.7 )
   END_RUNG
   RUNG wire#w1
      R_Coil( %DB60.DBX2.0 )
   END_RUNG
   RUNG wire#w1
      R_Coil( %DB60.DBX2.1 )
   END_RUNG
   RUNG wire#w1
      R_Coil( %DB60.DBX2.2 )
   END_RUNG
   RUNG wire#w1
      R_Coil( %DB60.DBX2.3 )
   END_RUNG
   RUNG wire#w1
      R_Coil( %DB60.DBX2.4 )
   END_RUNG
   RUNG wire#w1
      R_Coil( %DB60.DBX2.5 )
   END_RUNG
   RUNG wire#w1
      R_Coil( %DB60.DBX2.6 )
   END_RUNG